// TIA Portal project "ConveyorSystem2oo3" (V20)

(* hardware
DEVICE "S7-1500/ET200MP station_1"  S7-1500 station
   slot 0: "Rail_0"  Rack  6ES7 590-1***0-0AA0
   slot 1: "PLC_1"  CPU 1516-3 PN/DP  6ES7 516-3AP03-0AB0  V4.0
      slot 3: "CPU display_1"  6ES7591-1BA00-0AA0
      slot 32768: "PROFINET interface_1"  X1
         slot 32769: "Port_1"  X1 P1
         slot 32770: "Port_2"  X1 P2
      slot 33024: "PROFINET interface_2"  X2
         slot 33025: "Port_1"  X2 P1
      slot 33280: "DP interface_1"  X3
      slot 34817: "Virtual CP interface port_1"  Virtual CP interface port  Virtual CP interface port FW V4.0
DEVICE "HMI_1"  MTP1500 Unified Comfort
   slot 0: "HMI_1"  MTP1500 Unified Comfort  6AV2 128-3QB06-0AXx  20.0.0.0
   slot 1: "HMI_RT_1"  MTP1500 Unified Comfort  6AV2 128-3QB06-0AXx  20.0.0.0
   slot 5: "HMI_1.IE_CP_1"  PROFINET Interface  20.0.0.0
      slot 1: "PROFINET Interface_1"  PROFINET Interface
         slot 1: "Port_1"  Port
         slot 2: "Port_2"  Port
   slot 6: "HMI_1.IE_CP_2"  PROFINET Interface  20.0.0.0
      slot 1: "PROFINET Interface_GBit"  PROFINET Interface
         slot 1: "Port_1"  Port
*)

// ===== PLC "PLC_1"  CPU 1516-3 PN/DP =====

VAR_GLOBAL   // PLC tag table "Default tag table"
   "strobe" AT %Q0.0 : Bool;
   "data" AT %Q0.1 : Bool;
   "ultraVal" AT %I0.0 : Bool;
   "limitSwitchVal" AT %I0.1 : Bool;
   "relaySignal" AT %I0.3 : Bool;
   "testFunction" AT %M0.0 : Bool;
   "ackWire" AT %I0.4 : Bool;
   "faultReset" AT %M0.1 : Bool;
   "startCMD" AT %M0.2 : Bool;
   "stopCMD" AT %M0.3 : Bool;
   "servoPos" AT %MW0 : Int;
   "manualMode" AT %M0.4 : Bool;
   "moveServoHome" AT %M2.0 : Bool;
   "moveServoClear" AT %M2.1 : Bool;
   "conveyorToggle" AT %M2.2 : Bool;
END_VAR

TYPE "Fault-Log"
   STRUCT
      SensID : Int := -1;
      System : Int := -1;
   END_STRUCT;
END_TYPE

DATA_BLOCK "FaultLogs"   // DB1
{ S7_Optimized_Access := 'TRUE' }
VERSION : 0.1
   VAR
      Header : ArrayDBHeader;
      THIS : Array[0..19] of "Fault-Log";
   END_VAR
BEGIN
   Header.LowerBound := 0;
   Header.UpperBound := 19;
   Header.Elements := 20;
   Header.PaddedSize := 4;
   Header.ElementSize := 4;
END_DATA_BLOCK

DATA_BLOCK "TestFunctionality_DB"   // DB3
{ S7_Optimized_Access := 'TRUE' }
VERSION : 0.1
// stored: InstanceOfName TestFunctionality
"TestFunctionality"
BEGIN
END_DATA_BLOCK

DATA_BLOCK "AddFault_DB"   // DB4
{ S7_Optimized_Access := 'TRUE' }
VERSION : 0.1
// stored: InstanceOfName AddFault
"AddFault"
BEGIN
END_DATA_BLOCK

DATA_BLOCK "ManualController_DB"   // DB5
{ S7_Optimized_Access := 'TRUE' }
VERSION : 0.1
// stored: InstanceOfName ManualController
"ManualController"
BEGIN
END_DATA_BLOCK

DATA_BLOCK "ConveyerController_DB"   // DB6
{ S7_Optimized_Access := 'TRUE' }
VERSION : 0.1
// stored: InstanceOfName ConveyerController
"ConveyerController"
BEGIN
END_DATA_BLOCK

// folder: System blocks/Program resources

DATA_BLOCK "dataStrobeWireTON"   // DB2
{ S7_Optimized_Access := 'TRUE' }
AUTHOR : Simatic
FAMILY : IEC
NAME : IEC_TMR
VERSION : 1.0
// stored: InstanceOfName IEC_TIMER
"IEC_TIMER"
BEGIN
END_DATA_BLOCK

// folder: (top level)

FUNCTION_BLOCK "TestFunctionality"   // FB1, SCL
{ S7_Optimized_Access := 'TRUE' }
VERSION : 0.1
   VAR_OUTPUT
      faultID : Int;
      passed : Bool;
      fault : Bool;
   END_VAR
   VAR
      stateExternal : Int;
      stateInternal : Int;
      prevTestFunction : Bool;
      wireTONIN : Bool;
      excuted : Bool;
      ArduinoCOM : Int := -1;
   END_VAR
BEGIN
   IF #prevTestFunction = FALSE AND "testFunction" = TRUE THEN
       #stateExternal := 1;
       #stateInternal := 1;
       #passed := FALSE;
   END_IF;

   CASE #stateExternal OF
       1:
           CASE #stateInternal OF
               1:
                   "data" := TRUE;
                   "strobe" := TRUE;
                   #wireTONIN := TRUE;

                   "dataStrobeWireTON".TON(IN := #wireTONIN,
                                           PT := T#100ms);

                   IF "ackWire" = TRUE THEN
                       #excuted := TRUE;
                   END_IF;


                   IF "dataStrobeWireTON".Q = TRUE THEN
                       "data" := FALSE;
                       "strobe" := FALSE;
                       #wireTONIN := FALSE;
                       #stateInternal := 2;
                   END_IF;
               2:
                   IF #excuted = TRUE THEN
                       #ArduinoCOM := 1;
                   END_IF;

                   IF #excuted = FALSE THEN
                       #faultID := 5;
                       #fault := TRUE;
                       #stateInternal := 0;
                       #stateExternal := 0;
                       #ArduinoCOM := 0;

                   ELSIF BOOL_TO_INT("limitSwitchVal") + BOOL_TO_INT(NOT "ultraVal") = 2 THEN
                       #fault := FALSE;
                       #stateInternal := 3;

                   ELSIF BOOL_TO_INT("limitSwitchVal") + BOOL_TO_INT(NOT "ultraVal") = 0 THEN
                       #faultID := 4;
                       #fault := TRUE;

                   ELSIF "limitSwitchVal" = FALSE THEN
                       #faultID := 1;
                       #fault := TRUE;

                   ELSIF "ultraVal" = TRUE THEN
                       #faultID := 3;
                       #fault := TRUE;
                   END_IF;

               3:
                   "relaySignal" := TRUE;
                   #excuted := FALSE;
                   #stateInternal := 1;
                   #stateExternal := 2;
           END_CASE;


       2:
           "relaySignal" := FALSE;
           CASE #stateInternal OF
               1:
                   "data" := FALSE;
                   "strobe" := TRUE;
                   #wireTONIN := TRUE;

                   "dataStrobeWireTON".TON(IN := #wireTONIN,
                                           PT := T#100ms);

                   IF "ackWire" = TRUE THEN
                       #excuted := TRUE;
                   END_IF;


                   IF "dataStrobeWireTON".Q = TRUE THEN
                       "data" := FALSE;
                       "strobe" := FALSE;
                       #wireTONIN := FALSE;
                       #stateInternal := 2;
                   END_IF;
               2:
                   IF #excuted = FALSE THEN
                       #faultID := 5;
                       #fault := TRUE;
                       #stateInternal := 0;
                       #stateExternal := 0;

                   ELSIF BOOL_TO_INT(NOT "limitSwitchVal") + BOOL_TO_INT("ultraVal") = 2 THEN
                       #fault := FALSE;
                       #stateInternal := 3;

                   ELSIF BOOL_TO_INT(NOT "limitSwitchVal") + BOOL_TO_INT("ultraVal") = 0 THEN
                       #faultID := 4;
                       #fault := TRUE;

                   ELSIF "limitSwitchVal" = TRUE THEN
                       #faultID := 1;
                       #fault := TRUE;

                   ELSIF "ultraVal" = FALSE THEN
                       #faultID := 3;
                       #fault := TRUE;
                   END_IF;
               3:
                   #excuted := FALSE;
                   #stateInternal := 0;
                   #stateExternal := 0;
                   #passed := TRUE;
           END_CASE;
   END_CASE;
   #prevTestFunction := "testFunction";
END_FUNCTION_BLOCK

FUNCTION_BLOCK "AddFault"   // FB2, SCL
{ S7_Optimized_Access := 'TRUE' }
VERSION : 0.1
   VAR_INPUT
      faultTest : Bool;
      faultC : Bool;
      faultIDC : Int;
      faultIDTest : Int;
      faultIDM : Int;
      faultM : Bool;
   END_VAR
   VAR
      prevFaultTest : Bool := false;
      Index : Int := 0;
      prevFaultIDC : Int;
      prevFaultC : Bool;
      prevFaultIDTest : Int;
      latestFaultID : Int := -1;
      latestFaultSys : Int := -1;
      prevfaultIDM : Int;
      prevfaultM : Bool;
   END_VAR
BEGIN
   IF #prevFaultTest = FALSE AND #faultTest = TRUE OR NOT (#prevFaultIDTest = #faultIDTest) THEN
       "FaultLogs"."THIS"[#Index].SensID := #faultIDTest;
       "FaultLogs"."THIS"[#Index].System := 1;

       #latestFaultID := #faultIDTest;
       #latestFaultSys := 1;

       #Index := #Index + 1;

       IF #Index > 19 THEN
           #Index := 0;
       END_IF;
   END_IF;


   IF #prevfaultM = FALSE AND #faultM = TRUE OR NOT (#prevfaultIDM = #faultIDM) THEN
       "FaultLogs"."THIS"[#Index].SensID := #faultIDM;
       "FaultLogs"."THIS"[#Index].System := 2;

       #latestFaultID := #faultIDM;
       #latestFaultSys := 2;

       #Index := #Index + 1;

       IF #Index > 19 THEN
           #Index := 0;
       END_IF;
   END_IF;

   IF #prevFaultC = FALSE AND #faultC = TRUE OR NOT (#prevFaultIDC = #faultIDC) THEN
       "FaultLogs"."THIS"[#Index].SensID := #faultIDC;
       "FaultLogs"."THIS"[#Index].System := 2;

       #latestFaultID := #faultIDC;
       #latestFaultSys := 0;

       #Index := #Index + 1;

       IF #Index > 19 THEN
           #Index := 0;
       END_IF;
   END_IF;

   #prevFaultTest := #faultTest;
   #prevFaultIDTest := #faultIDTest;
   #prevFaultC := #faultC;
   #prevFaultIDC := #faultIDC;
   #prevfaultM := #faultM;
   #prevfaultIDM := #faultIDM;
END_FUNCTION_BLOCK

FUNCTION_BLOCK "ManualController"   // FB3, SCL
{ S7_Optimized_Access := 'TRUE' }
VERSION : 0.1
   VAR_OUTPUT
      fault : Bool;
      faultID : Int := -1;
   END_VAR
   VAR
      prevMoveHomeCMD : Bool;
      prevCloseCMD : Bool;
      prevconveyorSignal : Bool;
      state : Int;
      wireTONIN : Bool;
      excuted : Bool;
   END_VAR
BEGIN
   IF "manualMode" = TRUE THEN
       IF #prevMoveHomeCMD = FALSE AND "moveServoHome" = TRUE THEN
           CASE #state OF
               1:
                   "data" := TRUE;
                   "strobe" := TRUE;
                   #wireTONIN := TRUE;

                   "dataStrobeWireTON".TON(IN := #wireTONIN,
                                           PT := T#100ms);

                   IF "ackWire" = TRUE THEN
                       #excuted := TRUE;
                   END_IF;


                   IF "dataStrobeWireTON".Q = TRUE THEN
                       "data" := FALSE;
                       "strobe" := FALSE;
                       #wireTONIN := FALSE;
                       #state := 2;
                   END_IF;
               2:
                   IF #excuted = FALSE THEN
                       #faultID := 5;
                       #fault := TRUE;
                       #state := 0;

                   ELSIF BOOL_TO_INT("limitSwitchVal") + BOOL_TO_INT(NOT "ultraVal") = 2 THEN
                       #fault := FALSE;
                       #state := 3;

                   ELSIF BOOL_TO_INT("limitSwitchVal") + BOOL_TO_INT(NOT "ultraVal") = 0 THEN
                       #faultID := 4;
                       #fault := TRUE;
                       #state := 0;

                   ELSIF "limitSwitchVal" = FALSE THEN
                       #faultID := 1;
                       #fault := TRUE;
                       #state := 0;


                   ELSIF "ultraVal" = TRUE THEN
                       #faultID := 3;
                       #fault := TRUE;
                       #state := 0;

                   END_IF;
               3:
                   #excuted := FALSE;
                   #state := 0;
           END_CASE;
       END_IF;

       IF #prevCloseCMD = FALSE AND "moveServoHome" = TRUE THEN
           CASE #state OF
               1:
                   "data" := FALSE;
                   "strobe" := TRUE;
                   #wireTONIN := TRUE;

                   "dataStrobeWireTON".TON(IN := #wireTONIN,
                                           PT := T#100ms);

                   IF "ackWire" = TRUE THEN
                       #excuted := TRUE;
                   END_IF;


                   IF "dataStrobeWireTON".Q = TRUE THEN
                       "data" := FALSE;
                       "strobe" := FALSE;
                       #wireTONIN := FALSE;
                       #state := 2;
                   END_IF;
               2:
                   IF #excuted = FALSE THEN
                       #faultID := 5;
                       #fault := TRUE;
                       #state := 0;

                   ELSIF BOOL_TO_INT(NOT "limitSwitchVal") + BOOL_TO_INT("ultraVal") = 2 THEN
                       #fault := FALSE;
                       #state := 3;

                   ELSIF BOOL_TO_INT(NOT "limitSwitchVal") + BOOL_TO_INT("ultraVal") = 0 THEN
                       #faultID := 4;
                       #fault := TRUE;
                       #state := 0;

                   ELSIF "limitSwitchVal" = TRUE THEN
                       #faultID := 1;
                       #fault := TRUE;
                       #state := 0;


                   ELSIF "ultraVal" = FALSE THEN
                       #faultID := 3;
                       #fault := TRUE;
                       #state := 0;

                   END_IF;
               3:
                   #excuted := FALSE;
                   #state := 0;
           END_CASE;
       END_IF;

       IF #prevconveyorSignal = FALSE AND "conveyorToggle" = TRUE THEN
           "relaySignal" := NOT "relaySignal";
       END_IF;
   END_IF;
END_FUNCTION_BLOCK

FUNCTION_BLOCK "ConveyerController"   // FB5, SCL
{ S7_Optimized_Access := 'TRUE' }
VERSION : 0.1
   VAR_OUTPUT
      fault : Bool;
      faultID : Int;
   END_VAR
   VAR
      stateInternal : Int;
      stateExternal : Int;
      prevStartCMD : Bool;
      prevStopCMD : Bool;
      wireTONIN : Bool;
      excuted : Bool;
   END_VAR
BEGIN
   IF #prevStartCMD = FALSE AND "startCMD" = TRUE AND #stateInternal = 0 AND "manualMode" = FALSE THEN
       #stateExternal := 1;
       #stateInternal := 1;
   END_IF;

   IF #prevStopCMD = FALSE AND "stopCMD" = TRUE AND #stateInternal = 0 AND "manualMode" = FALSE THEN
       #stateExternal := 2;
       #stateInternal := 1;
   END_IF;


   CASE #stateExternal OF
       1:
           CASE #stateInternal OF
               1:
                   "data" := TRUE;
                   "strobe" := TRUE;
                   #wireTONIN := TRUE;

                   "dataStrobeWireTON".TON(IN := #wireTONIN,
                                           PT := T#100ms);

                   IF "ackWire" = TRUE THEN
                       #excuted := TRUE;
                   END_IF;


                   IF "dataStrobeWireTON".Q = TRUE THEN
                       "data" := FALSE;
                       "strobe" := FALSE;
                       #wireTONIN := FALSE;
                       #stateInternal := 2;
                   END_IF;
               2:
                   IF #excuted = FALSE THEN
                       #faultID := 5;
                       #fault := TRUE;
                       #stateInternal := 0;
                       #stateExternal := 0;

                   ELSIF BOOL_TO_INT("limitSwitchVal") + BOOL_TO_INT(NOT "ultraVal") = 2 THEN
                       #fault := FALSE;
                       #stateInternal := 3;

                   ELSIF BOOL_TO_INT("limitSwitchVal") + BOOL_TO_INT(NOT "ultraVal") = 0 THEN
                       #faultID := 4;
                       #fault := TRUE;
                       #stateInternal := 0;
                       #stateExternal := 0;


                   ELSIF "limitSwitchVal" = FALSE THEN
                       #faultID := 1;
                       #fault := TRUE;
                       #stateInternal := 0;
                       #stateExternal := 0;


                   ELSIF "ultraVal" = TRUE THEN
                       #faultID := 3;
                       #fault := TRUE;
                       #stateInternal := 0;
                       #stateExternal := 0;

                   END_IF;
               3:
                   "relaySignal" := TRUE;
                   #excuted := FALSE;
                   #stateInternal := 0;
                   #stateExternal := 0;
           END_CASE;


       2:
           "relaySignal" := FALSE;
           CASE #stateInternal OF
               1:
                   "data" := FALSE;
                   "strobe" := TRUE;
                   #wireTONIN := TRUE;

                   "dataStrobeWireTON".TON(IN := #wireTONIN,
                                           PT := T#100ms);

                   IF "ackWire" = TRUE THEN
                       #excuted := TRUE;
                   END_IF;


                   IF "dataStrobeWireTON".Q = TRUE THEN
                       "data" := FALSE;
                       "strobe" := FALSE;
                       #wireTONIN := FALSE;
                       #stateInternal := 2;
                   END_IF;
               2:
                   IF #excuted = FALSE THEN
                       #faultID := 5;
                       #fault := TRUE;
                       #stateInternal := 0;
                       #stateExternal := 0;

                   ELSIF BOOL_TO_INT(NOT "limitSwitchVal") + BOOL_TO_INT("ultraVal") = 2 THEN
                       #fault := FALSE;
                       #stateInternal := 3;

                   ELSIF BOOL_TO_INT(NOT "limitSwitchVal") + BOOL_TO_INT("ultraVal") = 0 THEN
                       #faultID := 4;
                       #fault := TRUE;
                       #stateInternal := 0;
                       #stateExternal := 0;

                   ELSIF "limitSwitchVal" = TRUE THEN
                       #faultID := 1;
                       #fault := TRUE;
                       #stateInternal := 0;
                       #stateExternal := 0;

                   ELSIF "ultraVal" = FALSE THEN
                       #faultID := 3;
                       #fault := TRUE;
                       #stateInternal := 0;
                       #stateExternal := 0;
                   END_IF;
               3:
                   #excuted := FALSE;
                   #stateInternal := 0;
                   #stateExternal := 0;
           END_CASE;
   END_CASE;

   #prevStopCMD := "stopCMD";
   #prevStartCMD := "startCMD";
END_FUNCTION_BLOCK

FUNCTION "ReadServoPos" : Void   // FC1, SCL
{ S7_Optimized_Access := 'TRUE' }
VERSION : 0.1
BEGIN
   IF BOOL_TO_INT("limitSwitchVal") + BOOL_TO_INT(NOT "ultraVal") = 2 THEN
       "servoPos" := 1;
   ELSIF BOOL_TO_INT(NOT "limitSwitchVal") + BOOL_TO_INT("ultraVal") = 2 THEN
       "servoPos" := 2;
   ELSE
       "servoPos" := 0;
   END_IF;
END_FUNCTION

ORGANIZATION_BLOCK "Main"   // OB1, SCL, ProgramCycle
TITLE = "Main Program Sweep (Cycle)"
{ S7_Optimized_Access := 'TRUE' }
VERSION : 0.1
   VAR_INPUT
      Initial_Call : Bool;   // Initial call of this OB
      Remanence : Bool;   // =True, if remanent data are available
   END_VAR
   VAR_TEMP
      faultIDtest : Int;
      testPassMain : Bool;
      faultTest : Bool;
      faultIDC : Int;
      faultC : Bool;
      faultIDM : Int;
      faultM : Bool;
   END_VAR
BEGIN
   "TestFunctionality_DB"(faultID=>#faultIDtest,
                          passed=>#testPassMain,
                          fault=>#faultTest);


   "ConveyerController_DB"(fault=>#faultC,
                           faultID=>#faultIDC);
   "AddFault_DB"(faultTest:=#faultTest,
                 faultC:=#faultC,
                 faultIDC:=#faultIDC,
                 faultIDTest:=#faultIDtest,
                 faultIDM:=#faultIDM,
                 faultM:=#faultM);




   "ManualController_DB"(fault=>#faultM,
                         faultID=>#faultIDM);


   "ReadServoPos"();
END_ORGANIZATION_BLOCK

(* ===== HMI "HMI_RT_1" =====
connection "HMI_Connection_1": ETHERNET, ILRT_S7_1500_OMS

HMI tags "Default tag table"
   "relaySignal" : Bool = PLC relaySignal AT %I0.3, T1s
   "ultraVal" : Bool = PLC ultraVal AT %I0.0, T1s
   "servoPos" : Int = PLC servoPos AT %MW0, T1s
   "limitSwitchVal" : Bool = PLC limitSwitchVal AT %I0.1, T1s
   "IRVal" : Bool = PLC IRVal AT %I0.2, T1s
   "TestFunctionality_DB_ArduinoCOM" : Int = PLC TestFunctionality_DB.ArduinoCOM, T1s
   "FaultLogs_THIS" : Array [0..19] of Fault-Log = PLC FaultLogs.THIS, T1s
   "FaultLogs_THIS{0}_SensID" : Int = PLC FaultLogs.THIS[0].SensID, T1s
   "AddFault_DB_Index" : Int = PLC AddFault_DB.Index, T1s
   "FIndex" : Int = PLC FIndex AT %MW2, T1s
   "AddFault_DB_latestFaultID" : Int = PLC AddFault_DB.latestFaultID, T1s
   "AddFault_DB_latestFaultSys" : Int = PLC AddFault_DB.latestFaultSys, T1s
   "startCMD" : Bool = PLC startCMD AT %M0.2, T1s
   "stopCMD" : Bool = PLC stopCMD AT %M0.3, T1s
   "manualMode" : Bool = PLC manualMode AT %M0.4, T1s
   "moveServoHome" : Bool = PLC moveServoHome AT %M2.0, T1s
   "moveServoClear" : Bool = PLC moveServoClear AT %M2.1, T1s
   "conveyorToggle" : Bool = PLC conveyorToggle AT %M2.2, T1s

text list "SystemTextList_ConfigErrorAlarmTextLibrary_1": 1 'NameService configuration error: Implicit deletion. Subelement instance @6%s@ must be deleted explicitly.'; 2 'NameService configuration error: Implicit deletion. Alias/Format/Unit instance @6%s@ must be deleted explicitly.'

text list "SystemTextList_ConfigErrorAlarmTextLibrary_2": 1 'EvDpManager::cleanupDeletedDatapoint - alert handler config is deleted implicitly for deleted datapoint, @3%s@'; 2 'EvDpManager::cleanupDeletedDatapoint - alert handler config is deleted implicitly but still has overrides, @3%s@'; 3 'EvDpManager::cleanupDeletedDatapoint - default value config is deleted implicitly for deleted datapoint, @3%s@'; 4 'EvDpManager::cleanupDeletedDatapoint - default value config is deleted implicitly but still has overrides, @3%s@'; 5 'EvDpManager::cleanupDeletedDatapoint - initial value config is deleted implicitly for deleted datapoint, @3%s@'; 6 'EvDpManager::cleanupDeletedDatapoint - initial value config is deleted implicitly but still has overrides, @3%s@'; 7 'EvDpManager::cleanupDeletedDatapoint - distribution config is deleted implicitly for deleted datapoint, @3%s@'; 8 'EvDpManager::cleanupDeletedDatapoint - distribution config is deleted implicitly but still has overrides, @3%s@'; 9 'EvDpManager::cleanupDeletedDatapoint - rangeCheck config is deleted implicitly for deleted datapoint, @3%s@'; 10 'EvDpManager::cleanupDeletedDatapoint - rangeCheck config is deleted implicitly but still has overrides, @3%s@'

text list "SystemTextList_ConfigErrorAlarmTextLibrary_3": 1 'The configured data point type was deleted, but a configured type is still defined for the node type: @3%s@.'; 2 'The configured data point node type was deleted in the data point type, but a configured type is still defined for the element: @3%s@.'

text list "SystemTextList_ConfigErrorAlarmTextLibrary_4": 2 'Cycles: @6%s@ does not exist'; 3 'Alarms: @6%s@ exists already'; 4 'Tags: Address @6%s@ was rejected'; 1 'Connections: @6%s@ does not exist'; 5 'Tags: Acquisition mode @6%s@ is not supported.'; 6 'Cycles: @6%s@ was deleted but associated tags exist.'; 7 'Connections: @6%s@ was deleted but associated tags exist.'; 8 'Tags: Tag @6%s@ was rejected.'; 9 'Tags: Tag @6%s@ has an invalid value.'; 0 'Connections: Connection to @6%s@ could not be established.'; 65638 'Connections: Connection to @6%s@ could not be established.'; 65639 'Connections: @6%s@ disconnected.'; 65640 'Connections: Connection to the HMI device @6%s@ is lost.'; 65641 'Connections: Connection to the PLC @6%s@ is lost.'; 65541 'Connections: Timeout while establishing the connection to @6%s@.'; 65542 'Connections: @6%s@ faulty.'; 65543 'Connections: Connection to the HMI device disconnected. Connection @5%s@ was changed.'; 65544 'Connections: Connection to the HMI device disconnected. Driver property was changed for connection @5%s@.'

text list "SystemTextList_ConfigErrorAlarmTextLibrary_5": 1 'Connections: Lifecycle monitoring cycle must be shorter than the response time.'; 2 'Connections: Cyclic services are configured but not supported by the target device.'; 3 'Connections: Change-controlled reading is configured but not supported by the target device.'; 4 'Tags: The address @6%s@ does not exist in the PLC.'; 5 'Tags: The default conversion type for the address @6%s@ could not be determined.'; 6 'Tags: Invalid conversion type'; 7 'Cycles: Invalid conversion type. Conversion is not supported at HmiCycle.'; 4096 'Connections: Version of the address @6%s@ is not supported.'; 4097 'Connections: PROFIBUS address is not supported.'; 4098 'Connections: Softbus address is not supported.'; 4099 'Connections: Address type @6%s@ is not supported.'; 4100 'Connections: Invalid connection name @6%s@. Access point is being ignored.'; 4101 'Connections: Routing is not supported. @6%s@ is not used.'; 4102 'Connections: Routing is not supported. @6%s@ is not used.'; 4103 'Connections: Invalid IP address @6%s@'; 4104 'Connections: Invalid Named Connection @6%s@. Valid format: >VMD</>connection<'; 4105 'Connections: Invalid Named Connection @6%s@. VMD connection name is too long. Only 24 characters are permitted.'; 4106 'Connections: Invalid Named Connection @6%s@. Connection name is too long. Only 32 characters are permitted.'; 4107 'Connections: Rack number @6%s@ is outside of the permitted range (0..7)'; 4108 'Connections: Invalid Named Connection @6%s@. Rack is ignored.'; 4109 'Connections: Slot number @6%s@ is outside of the permitted range (0..31)'; 4110 'Connections: Invalid Named Connection @6%s@. Slot is ignored.'; 4111 'Connection could not be established. Maximum number of available connections (@6%s@) has been exceeded.'; 4112 'Connection aborted. No sign of life in the last @4%s@ ms.'; 4113 'Connection could not be established - @4%s@'; 4114 'Connection could not be established. The address @6%s@ cannot be used.'; 4115 'Connection could not be established. Invalid address @6%s@'; 4116 'Connection could not be established - @4%s@'

text list "SystemTextList_ConfigErrorAlarmTextLibrary_6": 1 'Connection could not be established. Application instance certificate is not configured.'; 2 'Connection could not be established. Server has rejected the client certificate. OPC UA status code @4%s@.'; 3 'Connection could not be established. Internal problem in the certificate store. OPC UA status code @4%s@'; 4 'Connection could not be established. Application instance certificate could not be loaded. OPC UA status code @4%s@'; 5 'Connection could not be established. Server has not provided a certificate. @4%s@'; 6 'Connection could not be established. Validation of server certificate has failed. OPC UA status code @4%s@.'; 7 'Connection was closed. Error during alarm synchronization. OPC UA status code @4%s@.'; 8 'Connection was closed. Alarm/event subscription has failed. The number of operations on the server has been exceeded.'; 9 'Connection was closed. Alarm/event subscription has failed. The number of alarm/event subscriptions on the server has been exceeded.'; 10 'Connection could not be established. Server reports a license problem. OPC UA status code @4%s@.'; 11 'Connection could not be established. Maximum number of server sessions has been exceeded.'; 12 'Connection could not be established. Safety configuration is inconsistent. @4%s@'; 13 'Connection could not be established. The address @4%s@ cannot be used.'; 14 'Connection could not be established. OPC UA status code @4%s@'; 15 'Connection aborted. OPC UA server was stopped.'; 16 'Connection aborted. No sign of life in the last @4%s@ ms.'; 17 'Connection was closed. OPC UA server maintenance.'; 18 'Connection could not be established. Invalid configuration of the authentication mode - @4%s@'; 19 'Connection could not be established. User could not be authenticated. OPC UA status code @4%s@'; 20 'Connection could not be established. Server does not permit anonymous connection. OPC UA status code @4%s@'; 21 'Connection could not be established. Certificate problem: Error when writing the safety-relevant data to @4%s@.'; 22 'Connection could not be established. Certificate problem: Unexpected file in the folder @4%s@ cannot be removed.'; 23 'Connection could not be established. User could not be authenticated. No user or password configured.'; 24 'Connection could not be established. Unexpected length of the server certificate. @4%s@'; 25 'Connection could not be established. @4%s@ is empty.'; 26 'Connection could not be established. @4%s@ has an unexpected format.'; 27 'Connection could not be established. Server endpoints cannot be read. OPC UA status code @4%s@'; 28 'Connection could not be established. No server endpoints were found. @4%s@'; 29 'Connection could not be established. Application instance certificate could not be found.'; 30 'Connection could not be established. Unexpected format of the certificate @4%s@.'; 31 'Connection could not be established. Unexpected format of the certificate block list @4%s@.'; 32 'Connection could not be established. User could not be authenticated. An encryption detail is invalid. @4%s@'; 34 'Connection could not be established. - The configured non-transparent redundancy mode @4%s@ is not supported.'; 101 'Tags: Address @6%s@ does not exist on the server.'; 103 'Tags: Address @6%s@ cannot be accessed.'; 104 'Tags: Acquisition mode is not supported for address @6%s@.'; 201 'Alarms: Address @6%s@ does not exist on the server.'; 202 'Alarms: Address @6%s@ cannot be used. The specified range filter is not an OPC UA Event Notifier.'; 203 'Alarms: Address @6%s@ cannot be used. The specified range filter does not exist on the server.'; 204 'Alarms: Address @6%s@ cannot be used because it is not an OPC UA event type.'; 205 'Alarms: Address @6%s@ cannot be used because the OPC UA condition type is not supported.'; 206 'Alarms: Address @6%s@ cannot be used because the event type does not exist on the server.'; 207 'Alarms: Acquisition type cannot be used for address @6%s@.'; 301 'Address @6%s@ cannot be used because the version number is missing.'; 302 'Address @6%s@ cannot be used because the version number is invalid.'; 303 'Address @6%s@ cannot be used because the number of '$' delimiters is invalid.'; 304 'Address @6%s@ cannot be used because the address type is invalid.'; 305 'Unsupported version @6%s@ of the address'; 401 'Unexpected OPC UA server response: @6%s@'

text list "SystemTextList_ConfigErrorAlarmTextLibrary_7": 1 'Messages: Invalid condition string for the alarm view @6%s@.'; 2 'Messages: Invalid status tag and bit for the alarm view @6%s@.'; 3 'Messages: Invalid control tag and bit for the alarm view @6%s@.'

text list "SystemTextList_ConfigErrorAlarmTextLibrary_8": 1 'Logs: Implicit deletion. Logging tag instance @6%s@ should be deleted but there are overloaded elements.'

text list "SystemTextList_ConfigErrorAlarmTextLibrary_9": 2 'Restart of the runtime is required.'; 3 'The correct storage medium must be ejected and inserted again.'

text list "SystemTextList_ConfigErrorAlarmTextLibrary_10": 1 'CDS cache - Cache folder cannot be created or reached: @6%s@'; 2 'LOC cache - Cache folder cannot be created or reached: @6%s@'

text list "SystemTextList_ConfigErrorAlarmTextLibrary_11": 2 'and synchronization will start automatically. Shutting down either of them during synchronization will not cause data loss.'; 3 'and synchronization is scheduled for: @5%Y-%m-%d %H:%M:%S@. Shutting down either of the computers will not cause data loss.'

text list "SystemTextList_RuntimeCollaborationFailureReason_1": 0 'Unknown error (@3%s@)'; 1 'The system is not running or there is a network problem'; 2 'Runtime is not started on the target device.'; 3 'The System ID does not match the expected System ID (@3%s@)'; 4 'The Collaboration name does not match the expected Collaboration name '@3%s@''; 5 'Wrong or unknown certificate'; 6 'Revoked certificate'; 7 'The time difference is too big.'; 8 'No common supported message version'; 9 'System ID (@3%s@) already exists'; 10 'System name (@3%s@) already exists'; 11 'ID/Name in local configuration for Runtime Collaboration already exists'

text list "SystemTextList_RedundancyRecoveryFailureReason_1": 0 'Data recovery request temporarily rejected until own recovery request has been responded to.'; 1 'Data recovery request rejected. Online backup running.'; 2 'Data recovery request rejected. Connection to the Event Manager is not established.'; 3 'Data recovery request temporarily rejected until delta activation is complete.'; 4 'Data recovery request temporarily rejected until alarms and tags are retentive.'; 5 'Data recovery request rejected. The obligatory file config.level.es is missing on the computer.'; 6 'Data recovery request was canceled by the Event Manager.'; 7 'The data synchronization between the devices has failed.'

text list "SystemTextList_S7PlusAlarmTextListCollection_1": 4096 'Connections: Connection to the PLC @4%s@ is lost'; 4097 'Connections: Connection to the HMI device @4%s@ is lost'; 4098 'Connections: Maximum number of connections exceeded - @4%s@'; 4099 'Out of resources on PLC - @4%s@'; 4100 'Legitimation failed, invalid or missing password - @4%s@'; 4101 'Request to open the connection failed - @4%s@'; 4102 'Connections: Cannot connect to PLC - @4%s@'; 4103 'Request to open the connection could not be sent'; 4104 'General certificate error for PLC - @4%s@'; 4105 'PLC certificate expired for PLC - @4%s@'; 4106 'PLC certificate is revoked for PLC - @4%s@'; 4107 'PLC certificate is untrustworthy. Manual trust is possible for - @4%s@'; 4108 'PLC certificate is untrustworthy. Manual trust is not possible for - @4%s@'

text list "SystemTextList_AllenBradleyEIPAlarmTextListCollection_7": 4096 'Connection lost on PLC side - @5%s@'; 4097 'Connection lost on HMI side - @5%s@'; 4098 'Maximum number of connections exceeded - @5%s@'; 4099 'Out of resources on PLC - @5%s@'; 4100 'Legitimation failed, invalid or missing password - @5%s@'; 4101 'Open request failed - @5%s@'; 4102 'Cannot connect to PLC - @5%s@'; 4103 'Open request could not be sent'; 4104 'root certificate expired for - @5%s@'; 4105 'PLC certificate untrusted for - @5%s@'

text list "SystemTextList_AllenBradleyDF1AlarmTextListCollection_9": 4096 'Connections: Connection to the PLC @5%s@ is lost'; 4097 'Connections: Connection to the HMI device @5%s@ is lost'; 4098 'Connections: Maximum number of connections exceeded - @5%s@'; 4099 'Out of resources on PLC - @5%s@'; 4100 'Legitimation failed, invalid or missing password - @5%s@'; 4101 'Request to open the connection failed - @5%s@'; 4102 'Connections: Cannot connect to PLC - @5%s@'; 4103 'Request to open the connection could not be sent'; 4104 'General certificate error for PLC - @5%s@'; 4105 'PLC certificate expired for PLC - @5%s@'; 4106 'PLC certificate is revoked for PLC - @5%s@'; 4107 'PLC certificate is untrustworthy. Manual trust is possible for - @5%s@'; 4108 'PLC certificate is untrustworthy. Manual trust is not possible for - @5%s@'

text list "SystemTextList_OmronEIPAlarmTextListCollection_6": 4096 'Connection lost on PLC side - @5%s@'; 4097 'Connection lost on HMI side - @5%s@'; 4098 'Maximum number of connections exceeded - @5%s@'; 4099 'Out of resources on PLC - @5%s@'; 4100 'Legitimation failed, invalid or missing password - @5%s@'; 4101 'Open request failed - @5%s@'; 4102 'Cannot connect to PLC - @5%s@'; 4103 'Open request could not be sent'; 4104 'root certificate expired for - @5%s@'; 4105 'PLC certificate untrusted for - @5%s@'

text list "SystemTextList_StdModbusTCPAlarmTextListCollection_5": 4096 'Connections: Connection to the PLC @5%s@ is lost'; 4097 'Connections: Connection to the HMI device @5%s@ is lost'; 4098 'Connections: Maximum number of connections exceeded - @5%s@'; 4099 'Out of resources on PLC - @5%s@'; 4100 'Legitimation failed, invalid or missing password - @5%s@'; 4101 'Request to open the connection failed - @5%s@'; 4102 'Connections: Cannot connect to PLC - @5%s@'; 4103 'Request to open the connection could not be sent'; 4104 'General certificate error for PLC - @5%s@'; 4105 'PLC certificate expired for PLC - @5%s@'; 4106 'PLC certificate is revoked for PLC - @5%s@'; 4107 'PLC certificate is untrustworthy. Manual trust is possible for - @5%s@'; 4108 'PLC certificate is untrustworthy. Manual trust is not possible for - @5%s@'

text list "SystemTextList_MitsubishiMCAlarmTextListCollection_4": 4096 'Connection lost on PLC side - @5%s@'; 4097 'Connection lost on HMI side - @5%s@'; 4098 'Maximum number of connections exceeded - @5%s@'; 4099 'Out of resources on PLC - @5%s@'; 4100 'Legitimation failed, invalid or missing password - @5%s@'; 4101 'Open request failed - @5%s@'; 4102 'Cannot connect to PLC - @5%s@'; 4103 'Open request could not be sent'; 4104 'root certificate expired for - @5%s@'; 4105 'PLC certificate untrusted for - @5%s@'

text list "SystemTextList_MitsubishiiQAlarmTextListCollection_3": 4096 'Connection lost on PLC side - @5%s@'; 4097 'Connection lost on HMI side - @5%s@'; 4098 'Maximum number of connections exceeded - @5%s@'; 4099 'Out of resources on PLC - @5%s@'; 4100 'Legitimation failed, invalid or missing password - @5%s@'; 4101 'Open request failed - @5%s@'; 4102 'Cannot connect to PLC - @5%s@'; 4103 'Open request could not be sent'; 4104 'root certificate expired for - @5%s@'; 4105 'PLC certificate untrusted for - @5%s@'

text list "SystemTextList_StdModbusRTUAlarmTextListCollection_8": 4096 'Connections: Connection to the PLC @5%s@ is lost'; 4097 'Connections: Connection to the HMI device @5%s@ is lost'; 4098 'Connections: Maximum number of connections exceeded - @5%s@'; 4099 'Out of resources on PLC - @5%s@'; 4100 'Legitimation failed, invalid or missing password - @5%s@'; 4101 'Request to open the connection failed - @5%s@'; 4102 'Connections: Cannot connect to PLC - @5%s@'; 4103 'Request to open the connection could not be sent'; 4104 'General certificate error for PLC - @5%s@'; 4105 'PLC certificate expired for PLC - @5%s@'; 4106 'PLC certificate is revoked for PLC - @5%s@'; 4107 'PLC certificate is untrustworthy. Manual trust is possible for - @5%s@'; 4108 'PLC certificate is untrustworthy. Manual trust is not possible for - @5%s@'

text list "SystemTextList_LogoAlarmTextListCollection_10": 4096 'Connections: Connection to the PLC @5%s@ is lost'; 4097 'Connections: Connection to the HMI device @5%s@ is lost'; 4098 'Connections: Maximum number of connections exceeded - @5%s@'; 4099 'Out of resources on PLC - @5%s@'; 4100 'Legitimation failed, invalid or missing password - @5%s@'; 4101 'Request to open the connection failed - @5%s@'; 4102 'Connections: Cannot connect to PLC - @5%s@'; 4103 'Request to open the connection could not be sent'; 4104 'General certificate error for PLC - @5%s@'; 4105 'PLC certificate expired for PLC - @5%s@'; 4106 'PLC certificate is revoked for PLC - @5%s@'; 4107 'PLC certificate is untrustworthy. Manual trust is possible for - @5%s@'; 4108 'PLC certificate is untrustworthy. Manual trust is not possible for - @5%s@'
*)